(* Logix 5000 project; controller NWGG 1756-L72 rev 35.12; software revision 35.00; part 13 of 19 *)
(* tags used below, declared in another part *)
   tmrWeightTest : TIMER;
   Weight_Seed : DINT;
   _103_TANK_42_RECEIVING_LEG_RUNNING : BOOL;
   _106_TANK_17_AUGER_RUNNING : BOOL;
   _107_TANKS_1THRU7_SOUTH_RUNNING : BOOL;
   _108_CENTER_BELT_RUNNING : BOOL;
   _109_RAW_RECEIVING_NORTH_BELT_RUNNING : BOOL;
   _110_TANK_16_AUGER_RUNNING : BOOL;
   _113_HIGHROLLER_TANKS_11TO15_RUNNING : BOOL;
   _114_TANKS_1THRU7_NORTH_RUNNING : BOOL;
   _11_TANK_41_42_HIGHROLLER_RUNNING : BOOL;
   _123_CLEAN_LEG_RUNNING : BOOL;
   _1_CLEAN_SEED_UPPER_BELT_RUNNING : BOOL;
   _35_JUMP_LEG_RUNNING : BOOL;
   _3_LOWER_TANK_CONVAYOR_24TO26_RUNNING : BOOL;
   _43_SCREENINGS_LEG_RUNNING : BOOL;
   _4_LOWER_TANK_CONVAYOR_21TO23_RUNNING : BOOL;
   _5_LOWER_CROSS_BELT_RUNNING : BOOL;
   _701_TRUCK_REVERSING_BELT_RUNNING : BOOL;
   _703_TREATER_JUMP_BELT_RUNNING : BOOL;
   _9_TREATER_CONVAYOR_RUNNING : BOOL;
   Analog : AI[160];
   Calibration_Max : REAL;
   InEUMax : REAL;
   TestTag : REAL;
   Truck_Scales : udt_Truck_Scale[2];
(* MainProgram, continued *)

ROUTINE Totals   (* function block diagram *)
   SHEET 1
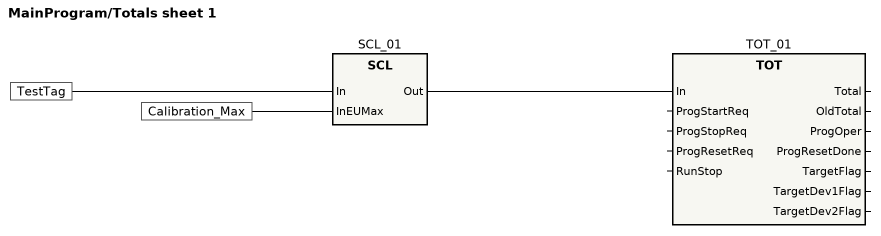
   SCL_01 : SCL(In := TestTag, InEUMax := Calibration_Max);
   TOT_01 : TOT(In := SCL_01.Out);   // unwired pins: ProgStartReq ProgStopReq ProgResetReq Total OldTotal ProgOper RunStop ProgResetDone TargetFlag TargetDev1Flag TargetDev2Flag
END_ROUTINE

ROUTINE VERIFACATION   (* ladder *)
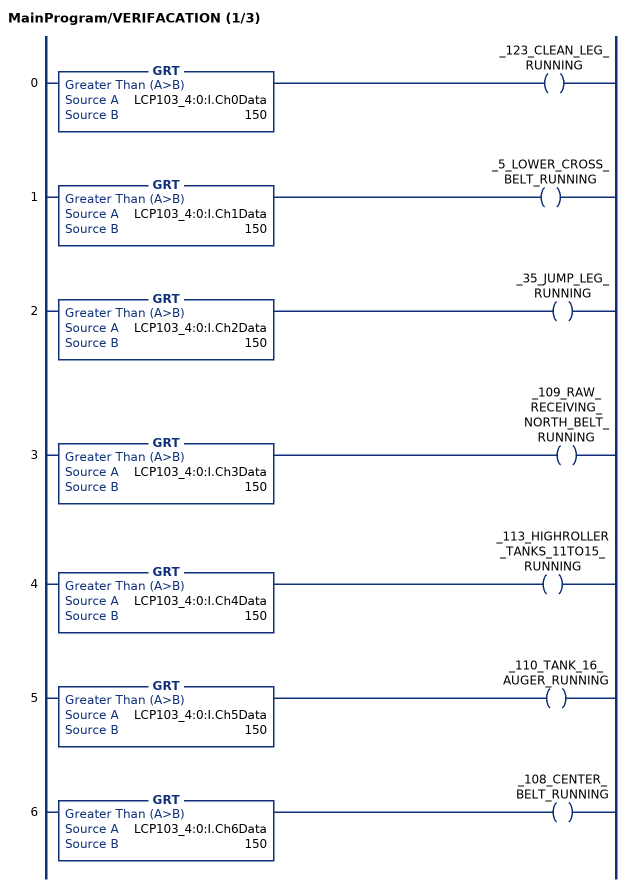
   0: GRT(LCP103_4:0:I.Ch0Data,150)OTE(_123_CLEAN_LEG_RUNNING);
   1: GRT(LCP103_4:0:I.Ch1Data,150)OTE(_5_LOWER_CROSS_BELT_RUNNING);
   2: GRT(LCP103_4:0:I.Ch2Data,150)OTE(_35_JUMP_LEG_RUNNING);
   3: GRT(LCP103_4:0:I.Ch3Data,150)OTE(_109_RAW_RECEIVING_NORTH_BELT_RUNNING);
   4: GRT(LCP103_4:0:I.Ch4Data,150)OTE(_113_HIGHROLLER_TANKS_11TO15_RUNNING);
   5: GRT(LCP103_4:0:I.Ch5Data,150)OTE(_110_TANK_16_AUGER_RUNNING);
   6: GRT(LCP103_4:0:I.Ch6Data,150)OTE(_108_CENTER_BELT_RUNNING);
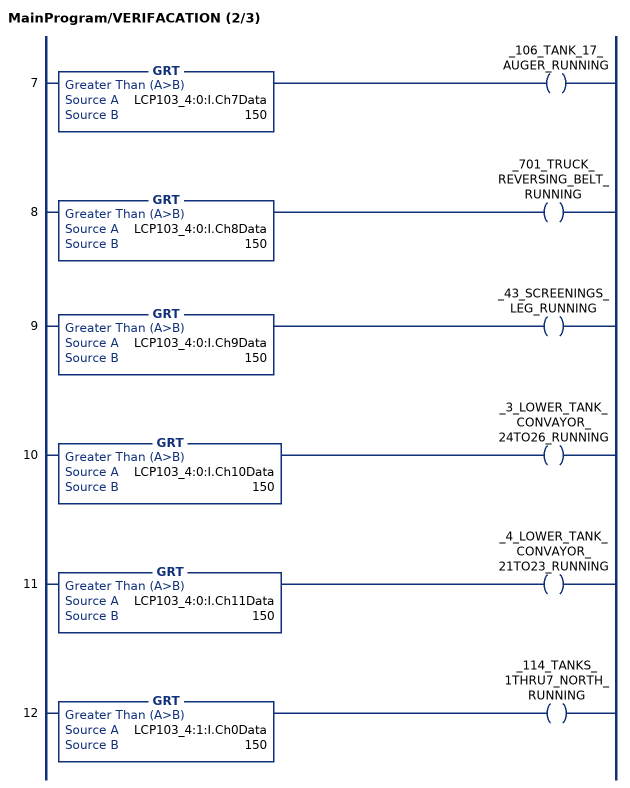
   7: GRT(LCP103_4:0:I.Ch7Data,150)OTE(_106_TANK_17_AUGER_RUNNING);
   8: GRT(LCP103_4:0:I.Ch8Data,150)OTE(_701_TRUCK_REVERSING_BELT_RUNNING);
   9: GRT(LCP103_4:0:I.Ch9Data,150)OTE(_43_SCREENINGS_LEG_RUNNING);
   10: GRT(LCP103_4:0:I.Ch10Data,150)OTE(_3_LOWER_TANK_CONVAYOR_24TO26_RUNNING);
   11: GRT(LCP103_4:0:I.Ch11Data,150)OTE(_4_LOWER_TANK_CONVAYOR_21TO23_RUNNING);
   12: GRT(LCP103_4:1:I.Ch0Data,150)OTE(_114_TANKS_1THRU7_NORTH_RUNNING);
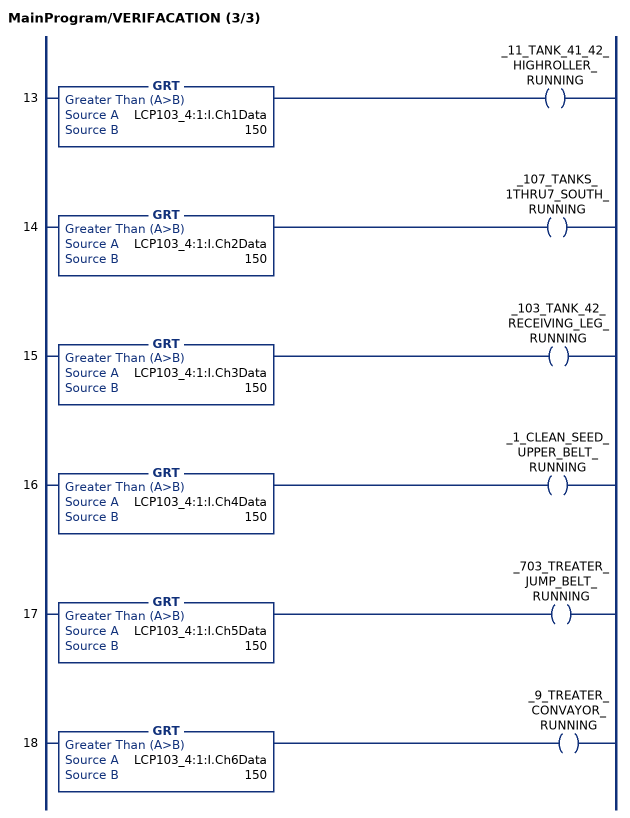
   13: GRT(LCP103_4:1:I.Ch1Data,150)OTE(_11_TANK_41_42_HIGHROLLER_RUNNING);
   14: GRT(LCP103_4:1:I.Ch2Data,150)OTE(_107_TANKS_1THRU7_SOUTH_RUNNING);
   15: GRT(LCP103_4:1:I.Ch3Data,150)OTE(_103_TANK_42_RECEIVING_LEG_RUNNING);
   16: GRT(LCP103_4:1:I.Ch4Data,150)OTE(_1_CLEAN_SEED_UPPER_BELT_RUNNING);
   17: GRT(LCP103_4:1:I.Ch5Data,150)OTE(_703_TREATER_JUMP_BELT_RUNNING);
   18: GRT(LCP103_4:1:I.Ch6Data,150)OTE(_9_TREATER_CONVAYOR_RUNNING);
END_ROUTINE

ROUTINE Weigh_Scales   (* ladder *)
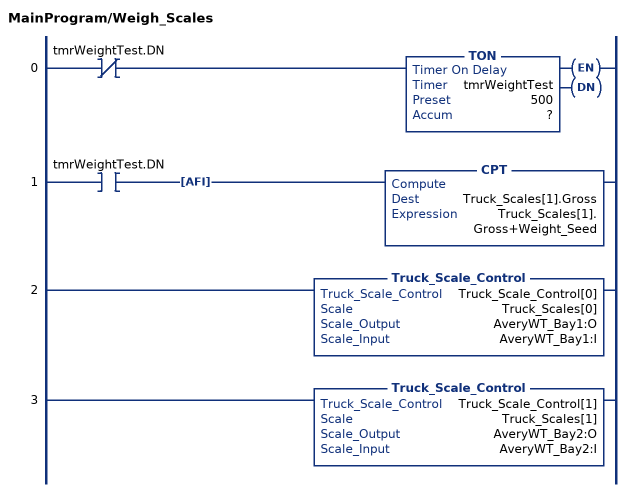
   0: XIO(tmrWeightTest.DN)TON(tmrWeightTest,?,?);
   1: XIC(tmrWeightTest.DN)AFI()CPT(Truck_Scales[1].Gross,Truck_Scales[1].Gross+Weight_Seed);
   2: Truck_Scale_Control(Truck_Scale_Control[0],Truck_Scales[0],AveryWT_Bay1:O,AveryWT_Bay1:I);
   3: Truck_Scale_Control(Truck_Scale_Control[1],Truck_Scales[1],AveryWT_Bay2:O,AveryWT_Bay2:I);
END_ROUTINE
END_PROGRAM

PROGRAM Scale   (* main routine MainRoutine *)
VAR
   ctlAddTime : CONTROL[2];
   ctrWtArray : COUNTER[2] := ([0].DN := 1, [1].DN := 1);
   Cur_Weight : REAL[2];
   Cur_Weight_Array_Idx : DINT := 16;
   Current_Gross : DINT[2];
   Current_Weight : REAL;
   Prev_Weight : REAL[2];
   Scale_Rate : REAL[2];
   Scale_Test_Rate_Mlt : DINT;
   ScaleIDX : DINT := 2;
   ShiftIDX : DINT := 20;
   TestRate : REAL[2];
   Time_Array : DINT[2,10] := ([0,0] := 9, [0,1] := 9, [0,2] := 10, [0,3] := 10, [0,4] := 8, [0,5] := 10, [0,6] := 9, [0,7] := 9, [0,8] := 9, [1,0] := 10, [1,1] := 9, [1,2] := 10, [1,3] := 10, [1,4] := 9, [1,5] := 10, [1,6] := 8, [1,7] := 10, [1,8] := 9);
   tmrRate : TIMER[2] := ([0].PRE := 1000, [0].ACC := 109, [0].EN := 1, [0].TT := 1, [1].PRE := 1000, [1].ACC := 126, [1].EN := 1, [1].TT := 1);
   tmrTestRate : TIMER[2] := ([1].ACC := 15, [1].EN := 1, [1].DN := 1);
   Total_Time : DINT[2];
   Weight_Array : REAL[2,40];
   Weight_Array_Idx : DINT[2] := ([0] := 14, [1] := 17);
   Weight_Array_Max : REAL[2];
   Weight_Sum : REAL[2];
END_VAR

ROUTINE AddWeights   (* ladder *)
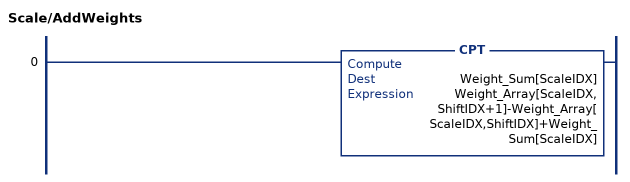
   0: CPT(Weight_Sum[ScaleIDX],Weight_Array[ScaleIDX,ShiftIDX+1]-Weight_Array[ScaleIDX,ShiftIDX]+Weight_Sum[ScaleIDX]);
END_ROUTINE

ROUTINE MainRoutine   (* ladder *)
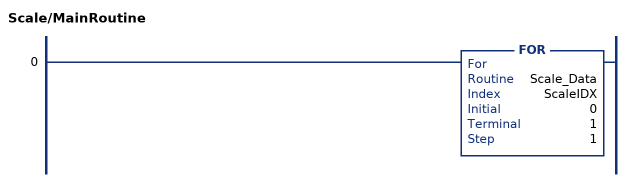
   0: FOR(Scale_Data,ScaleIDX,0,1,1);
END_ROUTINE

ROUTINE Scale_Data   (* ladder *)
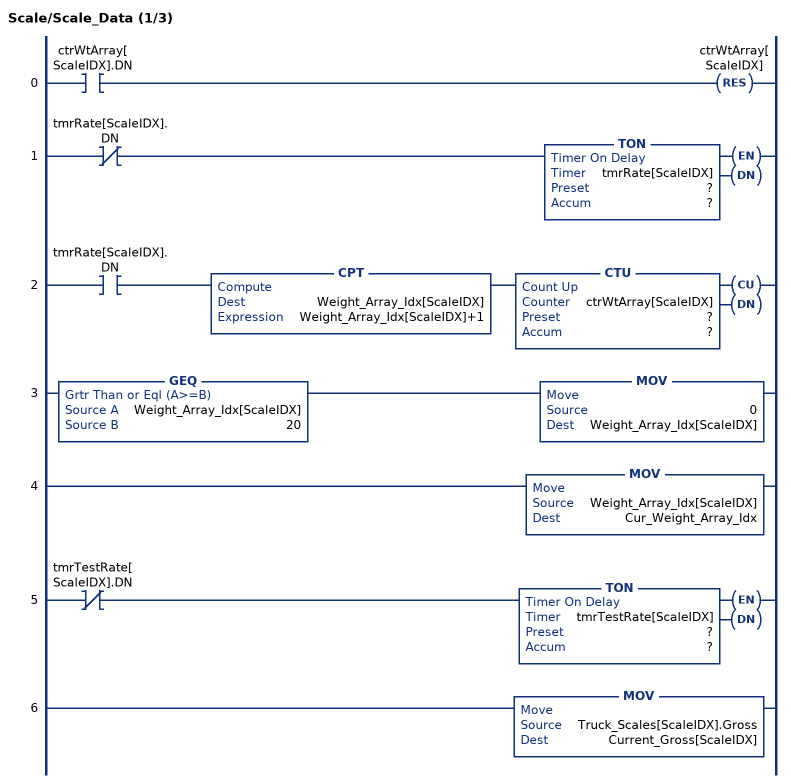
   0: XIC(ctrWtArray[ScaleIDX].DN)RES(ctrWtArray[ScaleIDX]);
   1: XIO(tmrRate[ScaleIDX].DN)TON(tmrRate[ScaleIDX],?,?);
   2: XIC(tmrRate[ScaleIDX].DN)CPT(Weight_Array_Idx[ScaleIDX],Weight_Array_Idx[ScaleIDX]+1)CTU(ctrWtArray[ScaleIDX],?,?);
   3: GEQ(Weight_Array_Idx[ScaleIDX],20)MOV(0,Weight_Array_Idx[ScaleIDX]);
   4: MOV(Weight_Array_Idx[ScaleIDX],Cur_Weight_Array_Idx);
   5: XIO(tmrTestRate[ScaleIDX].DN)TON(tmrTestRate[ScaleIDX],?,?);
   6: MOV(Truck_Scales[ScaleIDX].Gross,Current_Gross[ScaleIDX]);
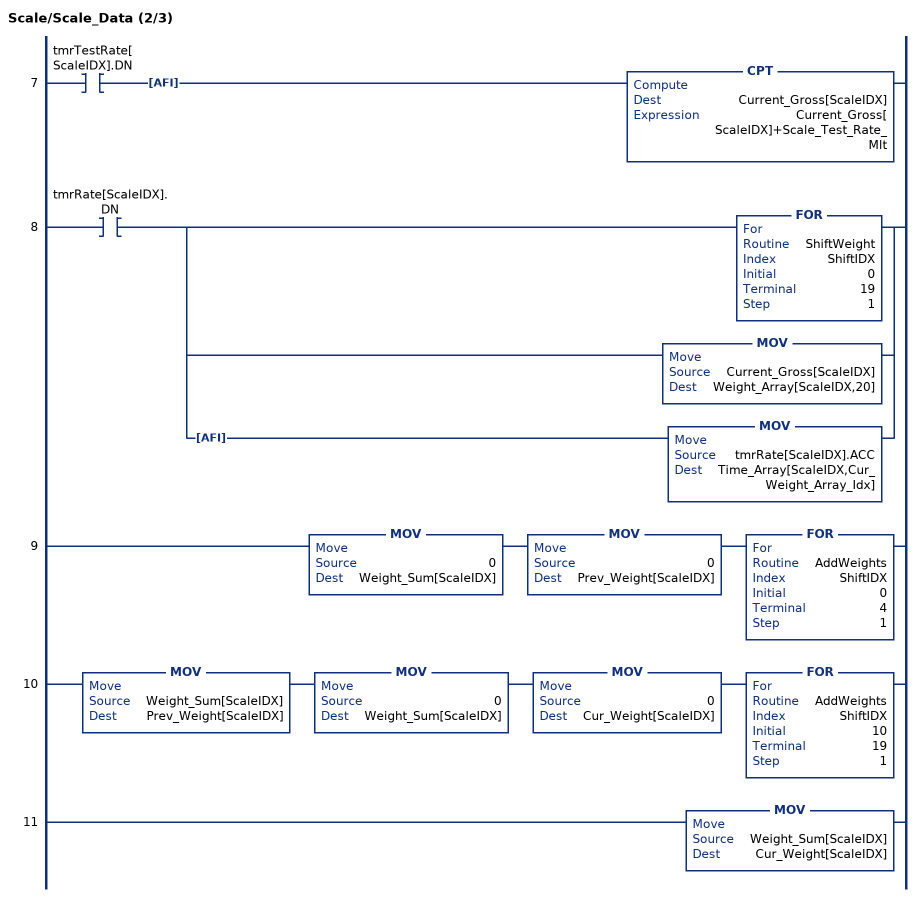
   7: XIC(tmrTestRate[ScaleIDX].DN)AFI()CPT(Current_Gross[ScaleIDX],Current_Gross[ScaleIDX]+Scale_Test_Rate_Mlt);
   8: XIC(tmrRate[ScaleIDX].DN)[FOR(ShiftWeight,ShiftIDX,0,19,1) ,MOV(Current_Gross[ScaleIDX],Weight_Array[ScaleIDX,20]) ,AFI() MOV(tmrRate[ScaleIDX].ACC,Time_Array[ScaleIDX,Cur_Weight_Array_Idx]) ];
   9: MOV(0,Weight_Sum[ScaleIDX])MOV(0,Prev_Weight[ScaleIDX])FOR(AddWeights,ShiftIDX,0,4,1);
   10: MOV(Weight_Sum[ScaleIDX],Prev_Weight[ScaleIDX])MOV(0,Weight_Sum[ScaleIDX])MOV(0,Cur_Weight[ScaleIDX])FOR(AddWeights,ShiftIDX,10,19,1);
   11: MOV(Weight_Sum[ScaleIDX],Cur_Weight[ScaleIDX]);
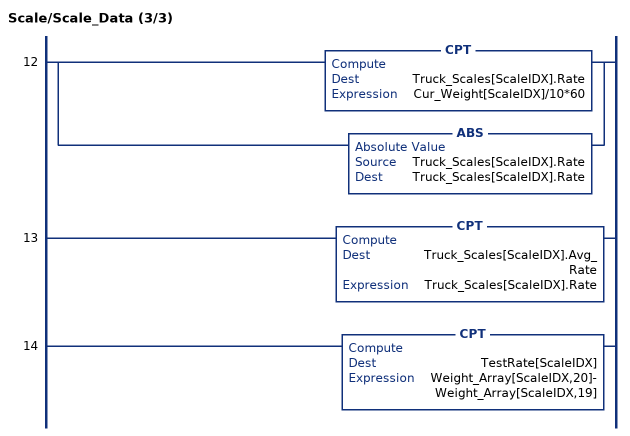
   12: [CPT(Truck_Scales[ScaleIDX].Rate,Cur_Weight[ScaleIDX]/10*60) ,ABS(Truck_Scales[ScaleIDX].Rate,Truck_Scales[ScaleIDX].Rate) ];
   13: CPT(Truck_Scales[ScaleIDX].Avg_Rate,Truck_Scales[ScaleIDX].Rate);
   14: CPT(TestRate[ScaleIDX],Weight_Array[ScaleIDX,20]-Weight_Array[ScaleIDX,19]);
END_ROUTINE

ROUTINE ShiftWeight   (* ladder *)
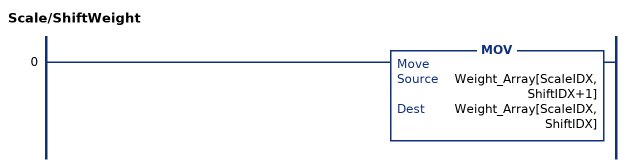
   0: MOV(Weight_Array[ScaleIDX,ShiftIDX+1],Weight_Array[ScaleIDX,ShiftIDX]);
END_ROUTINE
END_PROGRAM

PROGRAM SeedLoadoutMain   (* main routine MainRoutine *)
VAR
   Accept_Bin_Cal : BOOL;
   Air_Gates_Opened : BOOL;
   All_Stop : BOOL;
   ALM_Air_Gate_Failed_Open_Bin0 : ALARM_DIGITAL;
   ALM_Air_Gate_Failed_Open_Bin1 : ALARM_DIGITAL;
   ALM_Air_Gate_Failed_Open_Bin10 : ALARM_DIGITAL;
   ALM_Air_Gate_Failed_Open_Bin11 : ALARM_DIGITAL;
   ALM_Air_Gate_Failed_Open_Bin12 : ALARM_DIGITAL;
   ALM_Air_Gate_Failed_Open_Bin13 : ALARM_DIGITAL;
   ALM_Air_Gate_Failed_Open_Bin14 : ALARM_DIGITAL;
   ALM_Air_Gate_Failed_Open_Bin15 : ALARM_DIGITAL;
   ALM_Air_Gate_Failed_Open_Bin16 : ALARM_DIGITAL;
   ALM_Air_Gate_Failed_Open_Bin17 : ALARM_DIGITAL;
   ALM_Air_Gate_Failed_Open_Bin18 : ALARM_DIGITAL;
   ALM_Air_Gate_Failed_Open_Bin19 : ALARM_DIGITAL;
   ALM_Air_Gate_Failed_Open_Bin2 : ALARM_DIGITAL;
   ALM_Air_Gate_Failed_Open_Bin20 : ALARM_DIGITAL;
   ALM_Air_Gate_Failed_Open_Bin21 : ALARM_DIGITAL;
   ALM_Air_Gate_Failed_Open_Bin22 : ALARM_DIGITAL;
   ALM_Air_Gate_Failed_Open_Bin23 : ALARM_DIGITAL;
   ALM_Air_Gate_Failed_Open_Bin24 : ALARM_DIGITAL;
   ALM_Air_Gate_Failed_Open_Bin25 : ALARM_DIGITAL;
   ALM_Air_Gate_Failed_Open_Bin26 : ALARM_DIGITAL;
   ALM_Air_Gate_Failed_Open_Bin27 : ALARM_DIGITAL;
   ALM_Air_Gate_Failed_Open_Bin28 : ALARM_DIGITAL;
   ALM_Air_Gate_Failed_Open_Bin3 : ALARM_DIGITAL;
   ALM_Air_Gate_Failed_Open_Bin4 : ALARM_DIGITAL;
   ALM_Air_Gate_Failed_Open_Bin5 : ALARM_DIGITAL;
   ALM_Air_Gate_Failed_Open_Bin6 : ALARM_DIGITAL;
   ALM_Air_Gate_Failed_Open_Bin7 : ALARM_DIGITAL;
   ALM_Air_Gate_Failed_Open_Bin8 : ALARM_DIGITAL;
   ALM_Air_Gate_Failed_Open_Bin9 : ALARM_DIGITAL;
   ALM_K_Valve1_Treat_Failed : ALARM_DIGITAL;
   ALM_KValve0_Clean_Failed : ALARM_DIGITAL;
   ALM_KValve0_Treat_Failed : ALARM_DIGITAL;
   ALM_KValve1_Clean_Failed : ALARM_DIGITAL;
   ALM_NOT_USED : ALARM_DIGITAL;
   ALM_OVRAMP_Belt10 : ALARM_DIGITAL;
   ALM_OVRAMP_Belt11 : ALARM_DIGITAL;
   ALM_OVRAMP_Belt2 : ALARM_DIGITAL;
   ALM_OVRAMP_Belt3 : ALARM_DIGITAL;
   ALM_OVRAMP_Belt4 : ALARM_DIGITAL;
   ALM_OVRAMP_Belt5 : ALARM_DIGITAL;
   ALM_OVRAMP_Belt6 : ALARM_DIGITAL;
   ALM_OVRAMP_Belt7 : ALARM_DIGITAL;
   ALM_OVRAMP_Belt8 : ALARM_DIGITAL;
   ALM_OVRAMP_Belt9 : ALARM_DIGITAL;
   ALM_OVRAMP_CPLeg : ALARM_DIGITAL;
   ALM_PLUG_Belt1 : ALARM_DIGITAL;
   ALM_PLUG_Belt10 : ALARM_DIGITAL;
   ALM_PLUG_Belt11 : ALARM_DIGITAL;
   ALM_PLUG_Belt2 : ALARM_DIGITAL;
   ALM_PLUG_Belt3 : ALARM_DIGITAL;
   ALM_PLUG_Belt4 : ALARM_DIGITAL;
   ALM_PLUG_Belt5 : ALARM_DIGITAL;
   ALM_PLUG_Belt6 : ALARM_DIGITAL;
   ALM_PLUG_Belt7 : ALARM_DIGITAL;
   ALM_PLUG_Belt8 : ALARM_DIGITAL;
   ALM_PLUG_Belt9 : ALARM_DIGITAL;
   ALM_PLUG_CPLeg : ALARM_DIGITAL;
   ALM_SLP10_Belt1 : ALARM_DIGITAL;
   ALM_SLP10_Belt10 : ALARM_DIGITAL;
   ALM_SLP10_Belt11 : ALARM_DIGITAL;
   ALM_SLP10_Belt2 : ALARM_DIGITAL;
   ALM_SLP10_Belt3 : ALARM_DIGITAL;
   ALM_SLP10_Belt4 : ALARM_DIGITAL;
   ALM_SLP10_Belt5 : ALARM_DIGITAL;
   ALM_SLP10_Belt6 : ALARM_DIGITAL;
   ALM_SLP10_Belt7 : ALARM_DIGITAL;
   ALM_SLP10_Belt8 : ALARM_DIGITAL;
   ALM_SLP10_Belt9 : ALARM_DIGITAL;
   ALM_SLP10_CPLeg : ALARM_DIGITAL;
   ALM_SLP20_Belt1 : ALARM_DIGITAL;
   ALM_SLP20_Belt10 : ALARM_DIGITAL;
   ALM_SLP20_Belt11 : ALARM_DIGITAL;
   ALM_SLP20_Belt2 : ALARM_DIGITAL;
   ALM_SLP20_Belt3 : ALARM_DIGITAL;
   ALM_SLP20_Belt4 : ALARM_DIGITAL;
   ALM_SLP20_Belt5 : ALARM_DIGITAL;
   ALM_SLP20_Belt6 : ALARM_DIGITAL;
   ALM_SLP20_Belt7 : ALARM_DIGITAL;
   ALM_SLP20_Belt8 : ALARM_DIGITAL;
   ALM_SLP20_Belt9 : ALARM_DIGITAL;
   ALM_SLP20_CPLeg : ALARM_DIGITAL;
   ALM_WONT_START_Belt1 : ALARM_DIGITAL;
   ALM_WONT_START_Belt10 : ALARM_DIGITAL;
   ALM_WONT_START_Belt11 : ALARM_DIGITAL;
   ALM_WONT_START_Belt2 : ALARM_DIGITAL;
   ALM_WONT_START_Belt3 : ALARM_DIGITAL;
   ALM_WONT_START_Belt4 : ALARM_DIGITAL;
   ALM_WONT_START_Belt5 : ALARM_DIGITAL;
   ALM_WONT_START_Belt6 : ALARM_DIGITAL;
   ALM_WONT_START_Belt7 : ALARM_DIGITAL;
   ALM_WONT_START_Belt8 : ALARM_DIGITAL;
   ALM_WONT_START_Belt9 : ALARM_DIGITAL;
   ALM_WONT_START_CPLeg : ALARM_DIGITAL;
   Always_Off : BOOL;
   Andco_Auto_Mode : BOOL;
   Andco_Rate : DINT;
   Auto_Mode : BOOL := 1;
   Auto_Mode_ONS : BOOL;
   Auto_Start_Reversing_Belt_Fans : BOOL;
   Auto_Start_Treatment : BOOL;
   Auto_Stop_Clean : BOOL;
   Auto_Stop_Clean_Belt_11 : BOOL;
   Auto_Stop_Transfer : BOOL;
   Auto_Stop_Treat : BOOL;
   Available_For_Clean_Loadout : DINT := 536870911;
   Available_For_Treat_Loadout : DINT := 536870911;
   b3 : ALARM_DIGITAL;
   B_Offset : REAL;
   Batch_Status : DINT;
   BC_3_Belt_Required : BOOL;
   BC_9_Interlock : BOOL;
   Belt : udt_Motor[16] := ([0].Motor_Start.Auto_Stop_Delay := 5000, [1].Motor_Start.Auto_Stop_Delay := 5000, [1].Motor_Control.Spd_10_Pct := 1, [1].Motor_Control.Motor_Amps := -0.32500002, [1].Motor_Control.Motor_Batch_Ready := 1, [1].Motor_Control.Motor_Batch_Ready_Clean := 1, [1].Motor_Control.Motor_Batch_Ready_Treat := 1, [1].Motor_Control.Motor_Batch_Ready_Transfer := 1, [1].Motor_Config.Definition := 'Middle Concrete', [1].Motor_Config.Wind_Up_Time := 3000, [1].Motor_Config.Stop_At_SLP20 := 1, [1].Motor_Config.Stop_At_Max_Amps := 1, [1].Motor_Config.Max_Amps := 1000.0, [2].Motor_Start.Auto_Stop_Delay := 5000, [2].Motor_Control.Spd_10_Pct := 1, [2].Motor_Control.Motor_Amps := -0.4125, [2].Motor_Control.Motor_Batch_Ready := 1, [2].Motor_Control.Motor_Batch_Ready_Clean := 1, [2].Motor_Control.Motor_Batch_Ready_Treat := 1, [2].Motor_Control.Motor_Batch_Ready_Transfer := 1, [2].Motor_Config.Definition := 'North Concrete', [2].Motor_Config.Wind_Up_Time := 3000, [2].Motor_Config.Stop_At_SLP20 := 1, [3].Motor_Start.Auto_Stop_Delay := 5000, [3].Motor_Control.Spd_10_Pct := 1, [3].Motor_Control.Motor_Amps := -0.5125, [3].Motor_Control.Motor_Batch_Ready := 1, [3].Motor_Control.Motor_Batch_Ready_Clean := 1, [3].Motor_Control.Motor_Batch_Ready_Treat := 1, [3].Motor_Control.Motor_Batch_Ready_Transfer := 1, [3].Motor_Config.Definition := 'South Concrete', [3].Motor_Config.Wind_Up_Time := 3000, [3].Motor_Config.Stop_At_SLP20 := 1, [4].Motor_Start.Auto_Stop_Delay := 5000, [4].Motor_Control.Motor_Amps := -0.05285539, [4].Motor_Control.Motor_Batch_Ready := 1, [4].Motor_Control.Motor_Batch_Ready_Clean := 1, [4].Motor_Control.Motor_Batch_Ready_Treat := 1, [4].Motor_Control.Motor_Batch_Ready_Transfer := 1, [4].Motor_Config.Definition := 'Reversing', [4].Motor_Config.Wind_Up_Time := 6000, [4].Motor_Config.Stop_At_SLP20 := 1, [5].Motor_Start.Auto_Stop_Delay := 5000, [5].Motor_Control.Spd_10_Pct := 1, [5].Motor_Control.Motor_Amps := 0.018231237, [5].Motor_Control.Motor_Batch_Ready := 1, [5].Motor_Control.Motor_Batch_Ready_Clean := 1, [5].Motor_Control.Motor_Batch_Ready_Treat := 1, [5].Motor_Control.Motor_Batch_Ready_Transfer := 1, [5].Motor_Config.Definition := 'Treat Jump', [5].Motor_Config.Wind_Up_Time := 3000, [5].Motor_Config.Stop_At_SLP20 := 1, [6].Motor_Start.Auto_Stop_Delay := 5000, [6].Motor_Control.Spd_10_Pct := 1, [6].Motor_Control.Motor_Amps := 0.013243717, [6].Motor_Control.Motor_Batch_Ready := 1, [6].Motor_Control.Motor_Batch_Ready_Clean := 1, [6].Motor_Control.Motor_Batch_Ready_Treat := 1, [6].Motor_Control.Motor_Batch_Ready_Transfer := 1, [6].Motor_Config.Definition := 'Clean Jump',
        [6].Motor_Config.Wind_Up_Time := 3000, [6].Motor_Config.Stop_At_SLP20 := 1, [6].Motor_Config.Plugged_Sensor_Disabled := 1, [7].Motor_Start.Auto_Stop_Delay := 5000, [7].Motor_Control.Spd_10_Pct := 1, [7].Motor_Control.Motor_Amps := -0.23403546, [7].Motor_Control.Motor_Batch_Ready := 1, [7].Motor_Control.Motor_Batch_Ready_Clean := 1, [7].Motor_Control.Motor_Batch_Ready_Treat := 1, [7].Motor_Control.Motor_Batch_Ready_Transfer := 1, [7].Motor_Config.Definition := 'BC-9', [7].Motor_Config.Wind_Up_Time := 3000, [7].Motor_Config.Stop_At_SLP20 := 1, [7].Motor_Config.Plugged_Sensor_Disabled := 1, [8].Motor_Start.Auto_Stop_Delay := 5000, [8].Motor_Control.Spd_20_Pct := 1, [8].Motor_Control.Motor_Amps := 0.001667556, [8].Motor_Control.Motor_Batch_Ready := 1, [8].Motor_Control.Motor_Batch_Ready_Clean := 1, [8].Motor_Control.Motor_Batch_Ready_Treat := 1, [8].Motor_Control.Motor_Batch_Ready_Transfer := 1, [8].Motor_Config.Definition := 'BC-4', [8].Motor_Config.Wind_Up_Time := 3000, [8].Motor_Config.Speed_Sensor_Disabled := 1, [8].Motor_Config.Plugged_Sensor_Disabled := 1, [9].Motor_Start.Auto_Stop_Delay := 5000, [9].Motor_Control.Spd_20_Pct := 1, [9].Motor_Control.Motor_Amps := 0.033333335, [9].Motor_Control.Motor_Batch_Ready := 1, [9].Motor_Control.Motor_Batch_Ready_Clean := 1, [9].Motor_Control.Motor_Batch_Ready_Treat := 1, [9].Motor_Control.Motor_Batch_Ready_Transfer := 1, [9].Motor_Config.Definition := 'BC-3', [9].Motor_Config.Wind_Up_Time := 3000, [10].Motor_Start.Auto_Stop_Delay := 5000, [10].Motor_Control.Spd_20_Pct := 1, [10].Motor_Control.Motor_Amps := 0.016583197, [10].Motor_Control.Motor_Batch_Ready := 1, [10].Motor_Control.Motor_Batch_Ready_Clean := 1, [10].Motor_Control.Motor_Batch_Ready_Treat := 1, [10].Motor_Control.Motor_Batch_Ready_Transfer := 1, [10].Motor_Config.Definition := 'High Roller', [10].Motor_Config.Wind_Up_Time := 3000, [11].Motor_Start.Auto_Stop_Delay := 5000, [11].Motor_Control.Spd_20_Pct := 1, [11].Motor_Control.Motor_Amps := -0.008290774, [11].Motor_Control.Motor_Batch_Ready := 1, [11].Motor_Control.Motor_Batch_Ready_Clean := 1, [11].Motor_Control.Motor_Batch_Ready_Treat := 1, [11].Motor_Control.Motor_Batch_Ready_Transfer := 1, [11].Motor_Config.Definition := 'BC-5', [11].Motor_Config.Wind_Up_Time := 3000, [12].Motor_Start.Auto_Stop_Delay := 5000);
   Belt_Amps_Scale : SCALE[11];
   Belt_Gate_Leg_ON : BOOL;
   Belts_Ready : BOOL := 1;
   Belts_Running : BOOL;
   Bin_Cal : BOOL;
   Bin_Cal_IDX : DINT := -1;
   Bin_Calibration : BOOL;
   Bin_Clean_Pause : BOOL;
   Bin_Gate_Test : BOOL := 1;
   Bin_Loadout_Control : Loadout_Bin_Control[29] := ([0].Use_Bindicator := 1, [0].RawAnalogTag := 10270, [1].RawAnalogTag := 9993, [2].Use_Bindicator := 1, [2].RawAnalogTag := 8109, [3].RawAnalogTag := 3610, [4].RawAnalogTag := 7694, [5].RawAnalogTag := 5041, [6].RawAnalogTag := 9661, [7].RawAnalogTag := 9884, [8].RawAnalogTag := 10717, [9].RawAnalogTag := 9078, [10].RawAnalogTag := 8853, [11].RawAnalogTag := 9587, [12].RawAnalogTag := 7657, [13].RawAnalogTag := 9087, [14].RawAnalogTag := 9078, [15].RawAnalogTag := 8853, [16].Use_Bindicator := 1, [16].RawAnalogTag := 14748, [17].Use_Bindicator := 1, [17].RawAnalogTag := 15440, [18].Use_Bindicator := 1, [18].RawAnalogTag := 14244, [19].Use_Bindicator := 1, [19].RawAnalogTag := 13454, [20].Use_Bindicator := 1, [20].RawAnalogTag := 14460, [21].Use_Auger_Relay := 1, [21].Use_Bindicator := 1, [21].RawAnalogTag := 6343, [22].Use_Auger_Relay := 1, [22].Use_Bindicator := 1, [22].RawAnalogTag := 8758, [23].Use_Bindicator := 1, [23].RawAnalogTag := 15944, [24].Use_Bindicator := 1, [24].RawAnalogTag := 15184, [25].Use_Bindicator := 1, [25].RawAnalogTag := 15745, [26].Use_Bindicator := 1, [26].RawAnalogTag := 15279, [27].Use_Bindicator := 1, [27].RawAnalogTag := 14611, [28].Use_Bindicator := 1, [28].RawAnalogTag := 15145);
   Bin_Open_test : BOOL := 1;
   Bin_Transfer_Pause : BOOL;
   Bin_Treat_Pause : BOOL;
   Bin_Use_Index : DINT;
   Bin_Variety_Id : STRING[30] := ([0] := '823048', [1] := '823054', [2] := '823058', [3] := '823038', [4] := '823082', [5] := '823090', [6] := '823054', [7] := '823001', [9] := '873002', [10] := '873002', [11] := '873003', [12] := '823072', [16] := '823098', [17] := '843022', [19] := '822087', [20] := '803003', [21] := '823093', [22] := '843036', [23] := '843001', [24] := '843002', [25] := '843022', [26] := '803003', [27] := '823087', [28] := '803021');
   Bins_Rqd : BOOL;
   Blow_Out_Time : DINT;
   Blow_Out_Time_Remaining : REAL := -0.016;
   Blower_707_Running : BOOL;
   boolTransferTime : BOOL;
   Cal_Bin_Status : DINT;
   Cal_Done : BOOL;
   Calibrate_Mode : BOOL;
   Cancel_Bin_Config : BOOL;
   ckIDX : DINT := 29;
   Clean_Batch_Status : DINT;
   Clean_Bin_Gates_Opened : BOOL := 1;
   Clean_Interlock : BOOL;
   Clean_K_Relay_Not_Used : BOOL := 1;
   Clean_Load_Requested : BOOL;
   Clean_Scale_Target : DINT;
   Clean_Scale_Unavailable : BOOL;
   CleanHours : DINT;
   CleanMinuets : DINT;
   CleanSeconds : DINT;
   cntCleanTime : COUNTER := (PRE := 1);
   cntTest : COUNTER := (PRE := 100, ACC := 4);
   cntTransferTime : COUNTER := (PRE := 1);
   cntTreatTime : COUNTER := (PRE := 1);
   Concrete_Belts_Ready : BOOL;
   Concrete_Bin_Timing_Offset : DINT := 5;
   Concrete_Clean_Belts_Ready : BOOL;
   Concrete_Fan_Start : BOOL;
   Concrete_Leg : udt_Motor := (Motor_Start.Auto_Stop_Delay := 1, Motor_Control.Spd_20_Pct := 1, Motor_Control.Spd_10_Pct := 1, Motor_Control.Motor_Amps := -0.4625, Motor_Control.Motor_Batch_Ready_Clean := 1, Motor_Control.Motor_Batch_Ready_Treat := 1, Motor_Control.Motor_Batch_Ready_Transfer := 1, Motor_Config.Definition := 'CONCRETE LEG', Motor_Config.Wind_Up_Time := 4000, Motor_Config.Speed_Sensor_Disabled := 1, Motor_Config.Plugged_Sensor_Disabled := 1);
   Concrete_Leg_Interlock : BOOL;
   Concrete_Leg_Rqd : BOOL;
   Config_Bin_Name : STRING;
   Config_Cancel_Bin : BOOL := 1;
   Config_Class : STRING;
   Config_Clean_Delay_Start : REAL;
   Config_Clean_Delay_Stop : REAL;
   Config_Item_Number : STRING;
   Config_Name : STRING;
   Config_Pounds_Per_Inch : REAL;
   Config_Save_Bin : BOOL;
   Config_Treat_Delay_Start : REAL;
   Config_Treat_Delay_Stop : REAL;
   Configure_Clean_Delay : DINT := 36000;
   Configure_LoadoutBin : udt_Loadout_Bin := (Bin_Description := '9', Bin_Variety.Item_Number := '382010', Clean_Load_Delay_Start := 36000, Treat_Load_Delay_Start := 36000, Andco_Values.Raw_Position := 7, Andco_Values.Max_Position := 103, Andco_Values.Preact := 3, Andco_Values.Percent_Open := 0.067961164, Andco_Values.New_Pos := 9, Andco_Values.Width := 6.0);
   Configure_Treat_Delay_Start : DINT := 36000;
   ConfigureIndex : DINT := -1;
   ConfirmStop : BOOL;
   Current_Dist_List_IDX : DINT := 15;
   Current_Dist_Position : STRING := '10';
   Current_Longest_Time : DINT;
   Current_System_Msg_idx : DINT;
   Current_Transfer_Bin_From : BOOL[32];
   Current_Transfer_Bin_To : BOOL[32];
   DeltaX : REAL := -3028.0;
   DeltaY : REAL := -1000.0;
   Empty_String : STRING; {constant}
   Empty_Variety_ID : STRING := '0'; {constant}
   Finish_Treat_Ok : BOOL;
   FSC_Reverse : CONTROL;
   High_Roller_Belt_Bins_Required : BOOL;
   IDX : DINT := 29;
   Interlock_Not_Used : BOOL := 1;
   loa : ALARM_DIGITAL;
   Loadout_Bin : udt_Loadout_Bin[29] := ([0].Bin_Description := '3', [0].Bin_Variety.Item_Number := '823048', [0].Bin_Variety.Name := 'SEAHAWK CERTIFIED SPRING SWH', [0].Bin_Variety.Class := 'Certified', [0].Rate_Cal_Points[1].Andco_Position := 3631, [0].Rate_Cal_Points[1].Rate := 1000, [0].Rate_Cal_Points[2].Andco_Position := 6242, [0].Rate_Cal_Points[2].Rate := 2000, [0].Rate_Cal_Points[3].Andco_Position := 7451, [0].Rate_Cal_Points[3].Rate := 3000, [0].Rate_Cal_Points[4].Andco_Position := 9390, [0].Rate_Cal_Points[4].Rate := 4000, [0].Clean_Load_Delay_Start := 36050, [0].Treat_Load_Delay_Start := 29000, [0].Andco_Values.Cal_Status := 4, [0].Andco_Values.Raw_Position := 9707, [0].Andco_Values.Max_Position := 15761, [0].Andco_Values.Preact := 20, [0].Andco_Values.Percent_Open := 0.63870245, [0].Andco_Values.New_Pos := 1, [0].Andco_Values.Width := 6.0, [0].Andco_Values.Rate := 4163.4863, [0].Andco_Values.Pounds_Per_Inch := 65.0, [0].Andco_Values.New_Rate := 20.0, [0].Andco_Values.Analog := 1, [0].Andco_Values.Min_Position := 563, [0].Andco_Values.Length := 12.0, [0].Andco_Values.InchesOpen := 7.6644297, [0].Andco_Values.AnalogValue := 10270, [0].Clean_Load_Delay_Stop := 36050, [0].Treat_Load_Delay_Stop := 32000, [0].tmrStopDelay.EN := 1, [0].tmrStopDelay.TT := 1, [0].Available_For_Clean_Load := 1, [0].Available_For_Treat_Load := 1, [1].Bin_Description := '1', [1].Bin_Variety.Item_Number := '823054', [1].Bin_Variety.Name := 'RYAN CERTIFIED SPRING SWH', [1].Bin_Variety.Class := 'Certified', [1].Bin_Variety.Color[0].Color := 1, [1].Rate_Cal_Points[1].Andco_Position := 3454, [1].Rate_Cal_Points[1].Rate := 1000, [1].Rate_Cal_Points[2].Andco_Position := 5979, [1].Rate_Cal_Points[2].Rate := 2000, [1].Rate_Cal_Points[3].Andco_Position := 7870, [1].Rate_Cal_Points[3].Rate := 3000, [1].Rate_Cal_Points[4].Andco_Position := 9015, [1].Rate_Cal_Points[4].Rate := 4000, [1].Clean_Load_Delay_Start := 36100, [1].Treat_Load_Delay_Start := 29000, [1].Andco_Values.Cal_Status := 2, [1].Andco_Values.Raw_Position := 9424, [1].Andco_Values.Max_Position := 14962, [1].Andco_Values.Preact := 20, [1].Andco_Values.Percent_Open := 0.65476274, [1].Andco_Values.New_Pos := 2, [1].Andco_Values.Width := 6.0, [1].Andco_Values.Rate := 4357.205, [1].Andco_Values.Pounds_Per_Inch := 86.6, [1].Andco_Values.New_Rate := 1.0,
        [1].Andco_Values.Analog := 1, [1].Andco_Values.Min_Position := 569, [1].Andco_Values.Length := 12.0, [1].Andco_Values.InchesOpen := 7.857153, [1].Andco_Values.AnalogValue := 9993, [1].Clean_Load_Delay_Stop := 35000, [1].Treat_Load_Delay_Stop := 35000, [1].tmrStartDelay.PRE := 3000, [1].tmrStopDelay.PRE := 1000, [1].tmrStopDelay.EN := 1, [1].tmrStopDelay.TT := 1, [1].StartDelayPre := 3000, [1].StopDelayPre := 1000, [1].Available_For_Clean_Load := 1, [1].Available_For_Treat_Load := 1, [2].Bin_Description := '11', [2].Bin_Variety.Item_Number := '823058', [2].Bin_Variety.Name := 'MPRESS CERTIFIED FALL SWH', [2].Bin_Variety.Class := 'Certified', [2].Bin_Variety.Color[0].Color := 1, [2].Rate_Cal_Points[1].Andco_Position := 3384, [2].Rate_Cal_Points[1].Rate := 1000, [2].Rate_Cal_Points[2].Andco_Position := 5322, [2].Rate_Cal_Points[2].Rate := 2000, [2].Rate_Cal_Points[3].Andco_Position := 6882, [2].Rate_Cal_Points[3].Rate := 3000, [2].Rate_Cal_Points[4].Andco_Position := 7544, [2].Rate_Cal_Points[4].Rate := 4000, [2].Clean_Load_Delay_Start := 36000, [2].Treat_Load_Delay_Start := 30000, [2].Andco_Values.Cal_Status := 2, [2].Andco_Values.Raw_Position := 7352, [2].Andco_Values.Max_Position := 13688, [2].Andco_Values.Preact := 20, [2].Andco_Values.Percent_Open := 0.5686002, [2].Andco_Values.New_Pos := 54, [2].Andco_Values.Width := 6.0, [2].Andco_Values.Rate := 3709.9697, [2].Andco_Values.Pounds_Per_Inch := 65.0, [2].Andco_Values.New_Rate := 4000.0, [2].Andco_Values.Analog := 1, [2].Andco_Values.Min_Position := 758, [2].Andco_Values.Length := 12.0, [2].Andco_Values.InchesOpen := 6.823202, [2].Andco_Values.AnalogValue := 8110, [2].Clean_Load_Delay_Stop := 36000, [2].Treat_Load_Delay_Stop := 33000, [2].tmrStopDelay.EN := 1, [2].tmrStopDelay.TT := 1, [2].Available_For_Clean_Load := 1, [2].Available_For_Treat_Load := 1, [3].Bin_Description := '9', [3].Bin_Variety.Item_Number := '823038', [3].Bin_Variety.Name := 'DRIVE CERTIFIED FALL SWH', [3].Bin_Variety.Class := 'Certified', [3].Bin_Variety.Color[0].Color := 1, [3].Rate_Cal_Points[1].Andco_Position := 1926, [3].Rate_Cal_Points[1].Rate := 1000, [3].Rate_Cal_Points[2].Andco_Position := 5008, [3].Rate_Cal_Points[2].Rate := 2000,
        [3].Rate_Cal_Points[3].Andco_Position := 6109, [3].Rate_Cal_Points[3].Rate := 3000, [3].Rate_Cal_Points[4].Andco_Position := 7052, [3].Rate_Cal_Points[4].Rate := 4000, [3].Clean_Load_Delay_Start := 36000, [3].Treat_Load_Delay_Start := 31000, [3].Andco_Values.Cal_Status := 2, [3].Andco_Values.Raw_Position := 3192, [3].Andco_Values.Max_Position := 13763, [3].Andco_Values.Preact := 20, [3].Andco_Values.Percent_Open := 0.23919071, [3].Andco_Values.Width := 6.0, [3].Andco_Values.Rate := 1410.7722, [3].Andco_Values.Pounds_Per_Inch := 65.0, [3].Andco_Values.Analog := 1, [3].Andco_Values.Min_Position := 418, [3].Andco_Values.Length := 12.0, [3].Andco_Values.InchesOpen := 2.8702886, [3].Andco_Values.AnalogValue := 3610, [3].Clean_Load_Delay_Stop := 36000, [3].Treat_Load_Delay_Stop := 34000, [3].tmrStopDelay.EN := 1, [3].tmrStopDelay.TT := 1, [3].Available_For_Clean_Load := 1, [3].Available_For_Treat_Load := 1, [4].Bin_Description := '5', [4].Bin_Variety.Item_Number := '823082', [4].Bin_Variety.Name := 'LCS DAGGER AX - 5235 COAXIUM CERTIFIED SWH', [4].Bin_Variety.Class := 'Certified', [4].Rate_Cal_Points[1].Andco_Position := 3130, [4].Rate_Cal_Points[1].Rate := 1000, [4].Rate_Cal_Points[2].Andco_Position := 5282, [4].Rate_Cal_Points[2].Rate := 2000, [4].Rate_Cal_Points[3].Andco_Position := 6505, [4].Rate_Cal_Points[3].Rate := 3000, [4].Rate_Cal_Points[4].Andco_Position := 7576, [4].Rate_Cal_Points[4].Rate := 4000, [4].Clean_Load_Delay_Start := 36000, [4].Treat_Load_Delay_Start := 30000, [4].Andco_Values.Cal_Status := 4, [4].Andco_Values.Raw_Position := 7436, [4].Andco_Values.Max_Position := 13094, [4].Andco_Values.Preact := 20, [4].Andco_Values.Tolerance := 1, [4].Andco_Values.Percent_Open := 0.5793082, [4].Andco_Values.New_Pos := 63, [4].Andco_Values.Width := 6.0, [4].Andco_Values.Rate := 3869.281, [4].Andco_Values.Pounds_Per_Inch := 65.0, [4].Andco_Values.New_Rate := 4000.0, [4].Andco_Values.Analog := 1, [4].Andco_Values.Min_Position := 258, [4].Andco_Values.Length := 12.0, [4].Andco_Values.InchesOpen := 6.9516983, [4].Andco_Values.AnalogValue := 7694, [4].Clean_Load_Delay_Stop := 36000, [4].Treat_Load_Delay_Stop := 33000, [4].tmrStopDelay.EN := 1, [4].tmrStopDelay.TT := 1, [4].Available_For_Clean_Load := 1,
        [4].Available_For_Treat_Load := 1, [5].Bin_Description := '4', [5].Bin_Variety.Item_Number := '823090', [5].Bin_Variety.Name := 'REAPER-0293 CERTIFIED SWH', [5].Bin_Variety.Class := 'Certified', [5].Bin_Variety.Color[0].Color := 1, [5].Rate_Cal_Points[1].Andco_Position := 2925, [5].Rate_Cal_Points[1].Rate := 1000, [5].Rate_Cal_Points[2].Andco_Position := 4802, [5].Rate_Cal_Points[2].Rate := 2000, [5].Rate_Cal_Points[3].Andco_Position := 6340, [5].Rate_Cal_Points[3].Rate := 3000, [5].Rate_Cal_Points[4].Andco_Position := 7786, [5].Rate_Cal_Points[4].Rate := 4000, [5].Clean_Load_Delay_Start := 38000, [5].Treat_Load_Delay_Start := 30000, [5].Andco_Values.Cal_Status := 4, [5].Andco_Values.Raw_Position := 4496, [5].Andco_Values.Max_Position := 12868, [5].Andco_Values.Preact := 20, [5].Andco_Values.Percent_Open := 0.36484623, [5].Andco_Values.Width := 6.0, [5].Andco_Values.Rate := 1836.9739, [5].Andco_Values.Pounds_Per_Inch := 65.0, [5].Andco_Values.Analog := 1, [5].Andco_Values.Min_Position := 545, [5].Andco_Values.Length := 12.0, [5].Andco_Values.InchesOpen := 4.3781548, [5].Andco_Values.AnalogValue := 5041, [5].Clean_Load_Delay_Stop := 60000, [5].Treat_Load_Delay_Stop := 34000, [5].tmrStartDelay.PRE := 1000, [5].tmrStopDelay.EN := 1, [5].tmrStopDelay.TT := 1, [5].StartDelayPre := 1000, [5].Available_For_Clean_Load := 1, [5].Available_For_Treat_Load := 1, [6].Bin_Description := '7', [6].Bin_Variety.Item_Number := '823054', [6].Bin_Variety.Name := 'RYAN CERTIFIED SPRING SWH', [6].Bin_Variety.Class := 'Certified', [6].Bin_Variety.Color[0].Color := 1, [6].Rate_Cal_Points[1].Andco_Position := 3297, [6].Rate_Cal_Points[1].Rate := 1000, [6].Rate_Cal_Points[2].Andco_Position := 5415, [6].Rate_Cal_Points[2].Rate := 2000, [6].Rate_Cal_Points[3].Andco_Position := 7178, [6].Rate_Cal_Points[3].Rate := 3000, [6].Rate_Cal_Points[4].Andco_Position := 9109, [6].Rate_Cal_Points[4].Rate := 4000, [6].Clean_Load_Delay_Start := 36000, [6].Treat_Load_Delay_Start := 30000, [6].Andco_Values.Cal_Status := 4, [6].Andco_Values.Raw_Position := 9035, [6].Andco_Values.Max_Position := 15835, [6].Andco_Values.Preact := 20, [6].Andco_Values.Percent_Open := 0.5940171, [6].Andco_Values.New_Pos := 67, [6].Andco_Values.Width := 6.0, [6].Andco_Values.Rate := 3961.6777,